(* Logix 5000 project; controller PLC_MCC1300_75F1 vendor 1 type 14 code 166 rev 32.11; software revision 32.04; part 29 of 83 *)
(* tags used below, declared in another part *)
   B3 : DINT[51];
   BENCH_BUZZER : ALIAS FOR O[74].12;
   C5 : COUNTER[51];
   CNV10_FLT : ALIAS FOR I[4].9;
   CNV11_FLT : ALIAS FOR I[4].10;
   CNV12_FLT : ALIAS FOR I[4].11;
   CNV1_FLT : ALIAS FOR I[4].0;
   CNV2_FLT : ALIAS FOR I[4].1;
   CNV3_FLT : ALIAS FOR I[4].2;
   CNV4_FLT : ALIAS FOR I[4].3;
   CNV5_FLT : ALIAS FOR I[4].4;
   CNV6_FLT : ALIAS FOR I[4].5;
   CNV7_FLT : ALIAS FOR I[4].6;
   CNV8_FLT : ALIAS FOR I[4].7;
   CNV9_FLT : ALIAS FOR I[4].8;
   CRUSH_ALL_ON : ALIAS FOR B3[0].0;
   DRV_STOP_DEB : ALIAS FOR T4[30].DN;
   FAST_BLINK : ALIAS FOR T4[2];
   Host_Read : INT[500];
   I : INT[128];   // Local Input Updates Input Slot 2
   M2_ALM_HORN_RLY : ALIAS FOR O[9].3;
   M2_BLUE_STKLTE : ALIAS FOR O[9].5;
   MMI_DATA : INT[64];   // MMI DATA For Fix 32
   MMI_FROM_MB : MESSAGE;
   MMI_TO_MB : MESSAGE;
   N130 : INT[8];
   N131 : INT[8];
   N14 : DINT[500];
   N72 : DINT[200];
   O : INT[128];
   REL_CRUSH_ALL_OFF : ALIAS FOR I[73].10;
   REL_CRUSH_ALL_ON : ALIAS FOR I[73].11;
   SLOW_BLINK : ALIAS FOR T4[0];
   T4 : TIMER[51];
   TD_ALM_HORN_RLY : ALIAS FOR O[21].3;
   TD_CS2S_Crush_All_Stacklight : ALIAS FOR O[70].15;   // Red Light mounted on the top of panel
   TD_DRV_FLT_LMP : ALIAS FOR O[21].0;
   TDN_CRUSH_ALL_OFF : ALIAS FOR I[44].12;
   TDN_CRUSH_ALL_ON : ALIAS FOR I[44].13;
   TDN_FLT : ALIAS FOR I[18].1;
   TDS_CRUSH_ALL_OFF : ALIAS FOR I[64].12;
   TDS_CRUSH_ALL_ON : ALIAS FOR I[64].13;
   TDS_FLT : ALIAS FOR I[18].2;
   TK_FLT : ALIAS FOR I[18].0;
   TMR_Power_Cycle : TIMER;
   xAlwaysOFF : BOOL;
(* MainProgram, continued *)

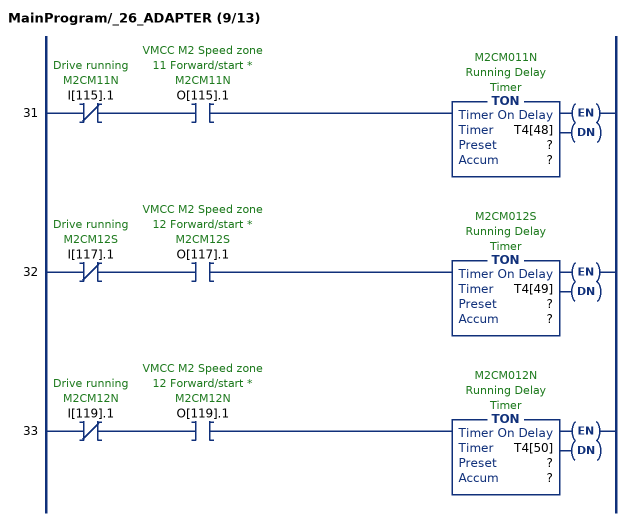
   31: XIO(I[115].1)XIC(O[115].1)TON(T4[48],?,?);
   32: XIO(I[117].1)XIC(O[117].1)TON(T4[49],?,?);
   33: XIO(I[119].1)XIC(O[119].1)TON(T4[50],?,?);
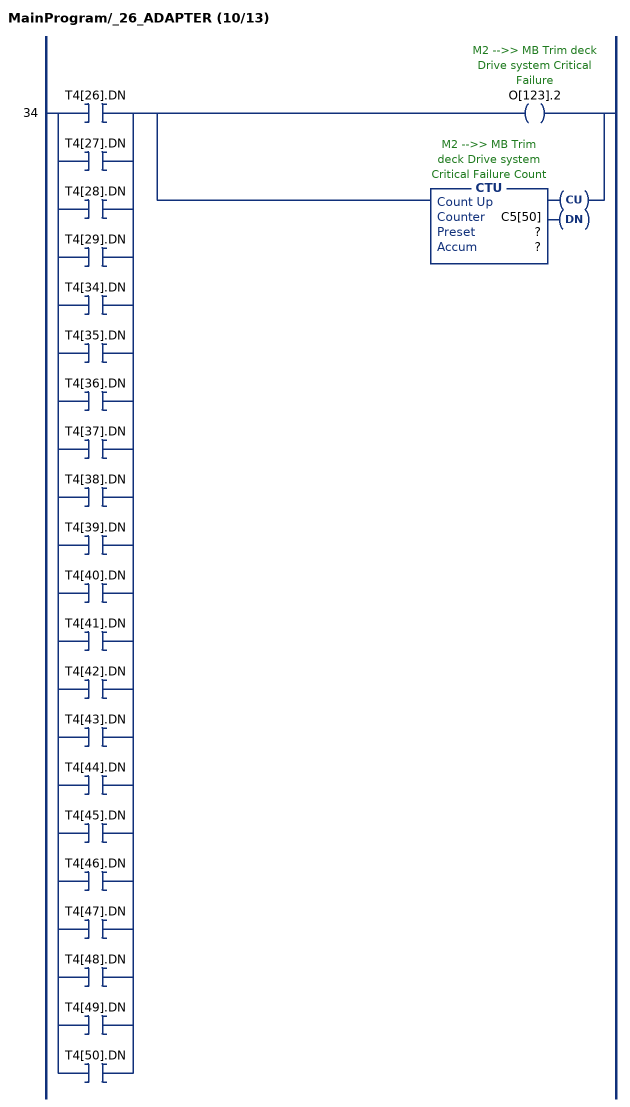
   34: [XIC(T4[26].DN) ,XIC(T4[27].DN) ,XIC(T4[28].DN) ,XIC(T4[29].DN) ,XIC(T4[34].DN) ,XIC(T4[35].DN) ,XIC(T4[36].DN) ,XIC(T4[37].DN) ,XIC(T4[38].DN) ,XIC(T4[39].DN) ,XIC(T4[40].DN) ,XIC(T4[41].DN) ,XIC(T4[42].DN) ,XIC(T4[43].DN) ,XIC(T4[44].DN) ,XIC(T4[45].DN) ,XIC(T4[46].DN) ,XIC(T4[47].DN) ,XIC(T4[48].DN) ,XIC(T4[49].DN) ,XIC(T4[50].DN) ][OTE(O[123].2) ,CTU(C5[50],?,?) ];
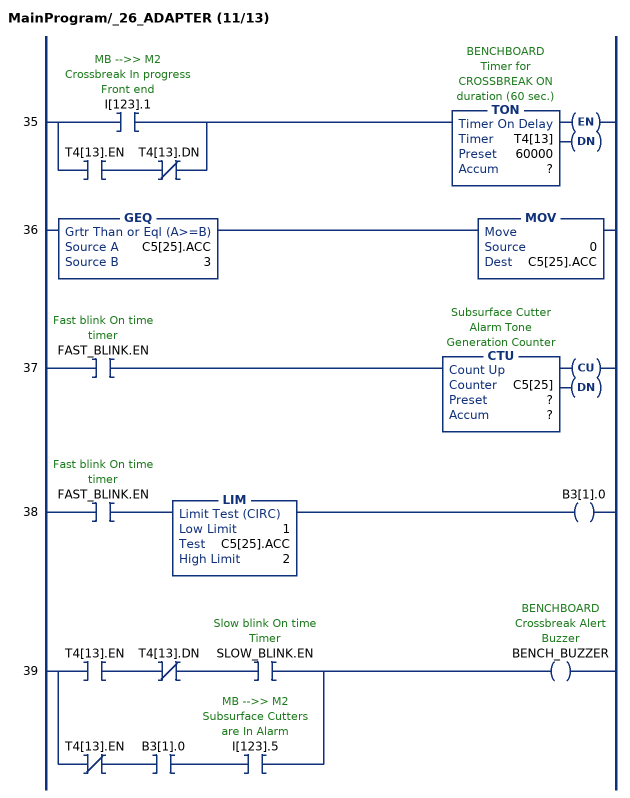
   35: [XIC(I[123].1) ,XIC(T4[13].EN) XIO(T4[13].DN) ]TON(T4[13],?,?);
   36: GEQ(C5[25].ACC,3)MOV(0,C5[25].ACC);
   37: XIC(FAST_BLINK.EN)CTU(C5[25],?,?);
   38: XIC(FAST_BLINK.EN)LIM(1,C5[25].ACC,2)OTE(B3[1].0);
   39: [XIC(T4[13].EN) XIO(T4[13].DN) XIC(SLOW_BLINK.EN) ,XIO(T4[13].EN) XIC(B3[1].0) XIC(I[123].5) ]OTE(BENCH_BUZZER);
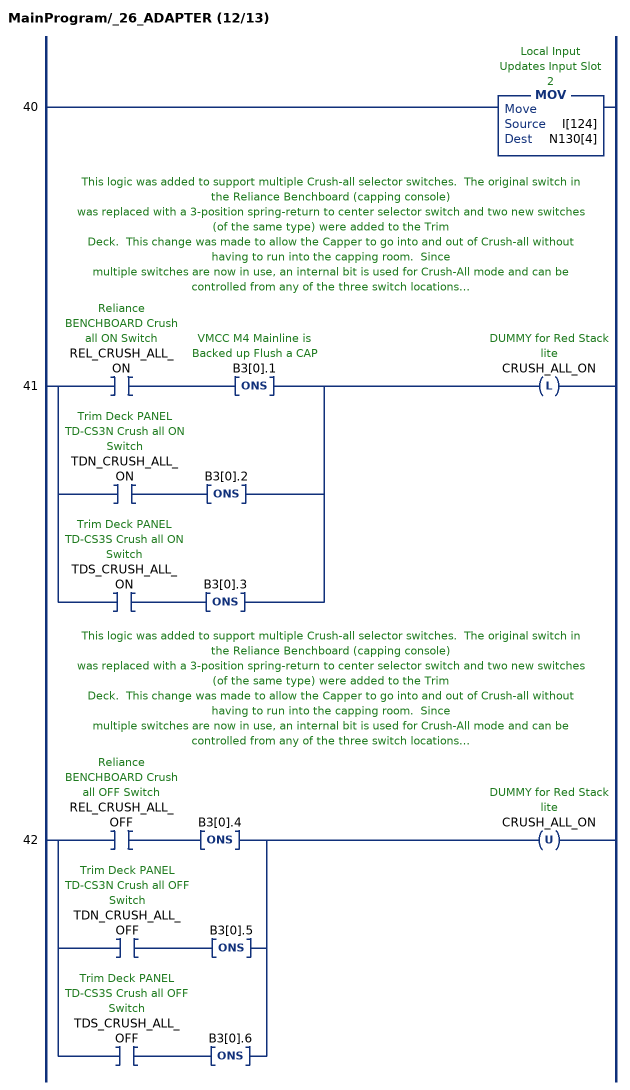
   40: MOV(I[124],N130[4]);
   // This logic was added to support multiple Crush-all selector switches.  The original switch in the Reliance Benchboard (capping console)
   // was replaced with a 3-position spring-return to center selector switch and two new switches (of the same type) were added to the Trim
   // Deck.  This change was made to allow the Capper to go into and out of Crush-all without having to run into the capping room.  Since
   // multiple switches are now in use, an internal bit is used for Crush-All mode and can be controlled from any of the three switch locations.
   // Note that one-shots [ONS] are used to keep a stuck-on selector switch contact from preventing the other two switches from operating
   // properly.  Also note that Latches and Unlatches are used (rather than a seal circuit) so that the system rides through power bumps properly
   // (i.e. Crush-all will stay in its current state, whether on or off, after a power bump).   DMK 10/21/02
   41: [XIC(REL_CRUSH_ALL_ON) ONS(B3[0].1) ,XIC(TDN_CRUSH_ALL_ON) ONS(B3[0].2) ,XIC(TDS_CRUSH_ALL_ON) ONS(B3[0].3) ]OTL(CRUSH_ALL_ON);
   // This logic was added to support multiple Crush-all selector switches.  The original switch in the Reliance Benchboard (capping console)
   // was replaced with a 3-position spring-return to center selector switch and two new switches (of the same type) were added to the Trim
   // Deck.  This change was made to allow the Capper to go into and out of Crush-all without having to run into the capping room.  Since
   // multiple switches are now in use, an internal bit is used for Crush-All mode and can be controlled from any of the three switch locations.
   // Note that one-shots [ONS] are used to keep a stuck-on selector switch contact from preventing the other two switches from operating
   // properly.  Also note that Latches and Unlatches are used (rather than a seal circuit) so that the system rides through power bumps properly
   // (i.e. Crush-all will stay in its current state, whether on or off, after a power bump).   DMK 10/21/02
   42: [XIC(REL_CRUSH_ALL_OFF) ONS(B3[0].4) ,XIC(TDN_CRUSH_ALL_OFF) ONS(B3[0].5) ,XIC(TDS_CRUSH_ALL_OFF) ONS(B3[0].6) ]OTU(CRUSH_ALL_ON);
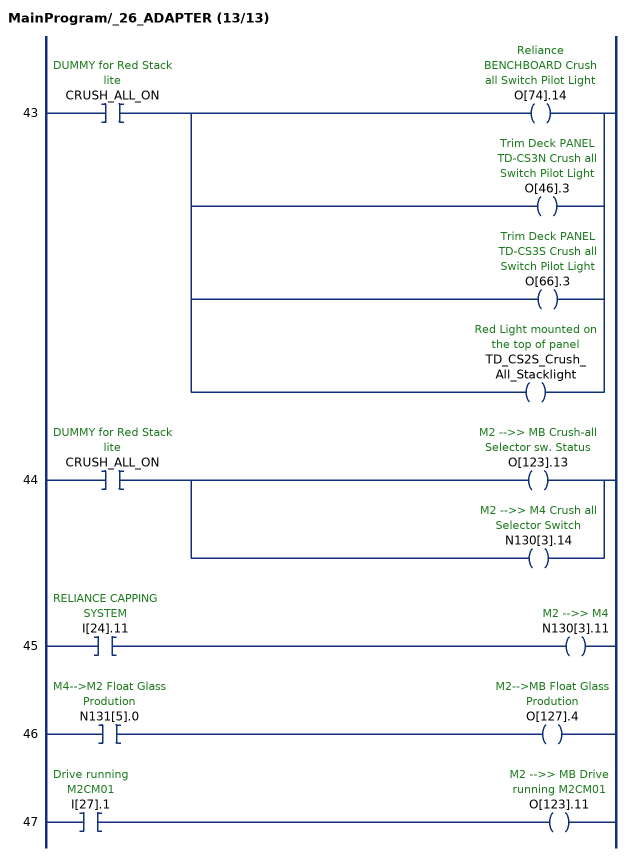
   43: XIC(CRUSH_ALL_ON)[OTE(O[74].14) ,OTE(O[46].3) ,OTE(O[66].3) ,OTE(TD_CS2S_Crush_All_Stacklight) ];
   44: XIC(CRUSH_ALL_ON)[OTE(O[123].13) ,OTE(N130[3].14) ];
   45: XIC(I[24].11)OTE(N130[3].11);
   46: XIC(N131[5].0)OTE(O[127].4);
   47: XIC(I[27].1)OTE(O[123].11);
END_ROUTINE

ROUTINE _2_MCP_A   (* ladder *)
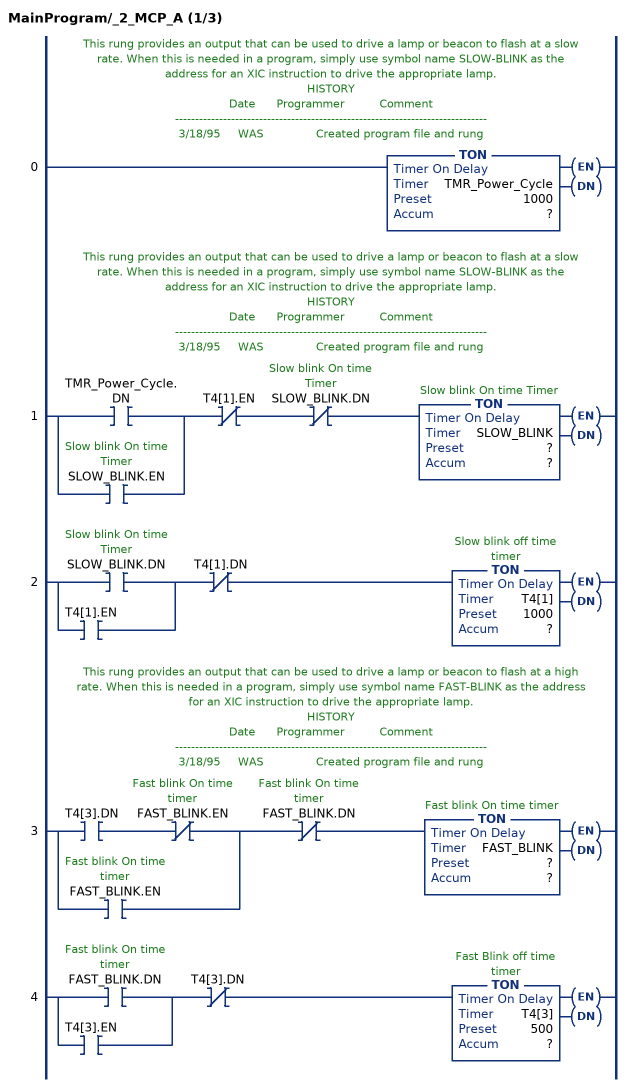
   // This rung provides an output that can be used to drive a lamp or beacon to flash at a slow rate. When this is needed in a program, simply use symbol name SLOW-BLINK as the address for an XIC instruction to drive the appropriate lamp.
   // HISTORY
   //             Date      Programmer          Comment
   // ------------------------------------------------------------------------------
   //             3/18/95     WAS               Created program file and rung
   0: TON(TMR_Power_Cycle,?,?);
   // This rung provides an output that can be used to drive a lamp or beacon to flash at a slow rate. When this is needed in a program, simply use symbol name SLOW-BLINK as the address for an XIC instruction to drive the appropriate lamp.
   // HISTORY
   //             Date      Programmer          Comment
   // ------------------------------------------------------------------------------
   //             3/18/95     WAS               Created program file and rung
   1: [XIC(TMR_Power_Cycle.DN) ,XIC(SLOW_BLINK.EN) ]XIO(T4[1].EN)XIO(SLOW_BLINK.DN)TON(SLOW_BLINK,?,?);
   2: [XIC(SLOW_BLINK.DN) ,XIC(T4[1].EN) ]XIO(T4[1].DN)TON(T4[1],?,?);
   // This rung provides an output that can be used to drive a lamp or beacon to flash at a high rate. When this is needed in a program, simply use symbol name FAST-BLINK as the address for an XIC instruction to drive the appropriate lamp.
   // HISTORY
   //             Date      Programmer          Comment
   // ------------------------------------------------------------------------------
   //             3/18/95     WAS               Created program file and rung
   3: [XIC(T4[3].DN) XIO(FAST_BLINK.EN) ,XIC(FAST_BLINK.EN) ]XIO(FAST_BLINK.DN)TON(FAST_BLINK,?,?);
   4: [XIC(FAST_BLINK.DN) ,XIC(T4[3].EN) ]XIO(T4[3].DN)TON(T4[3],?,?);
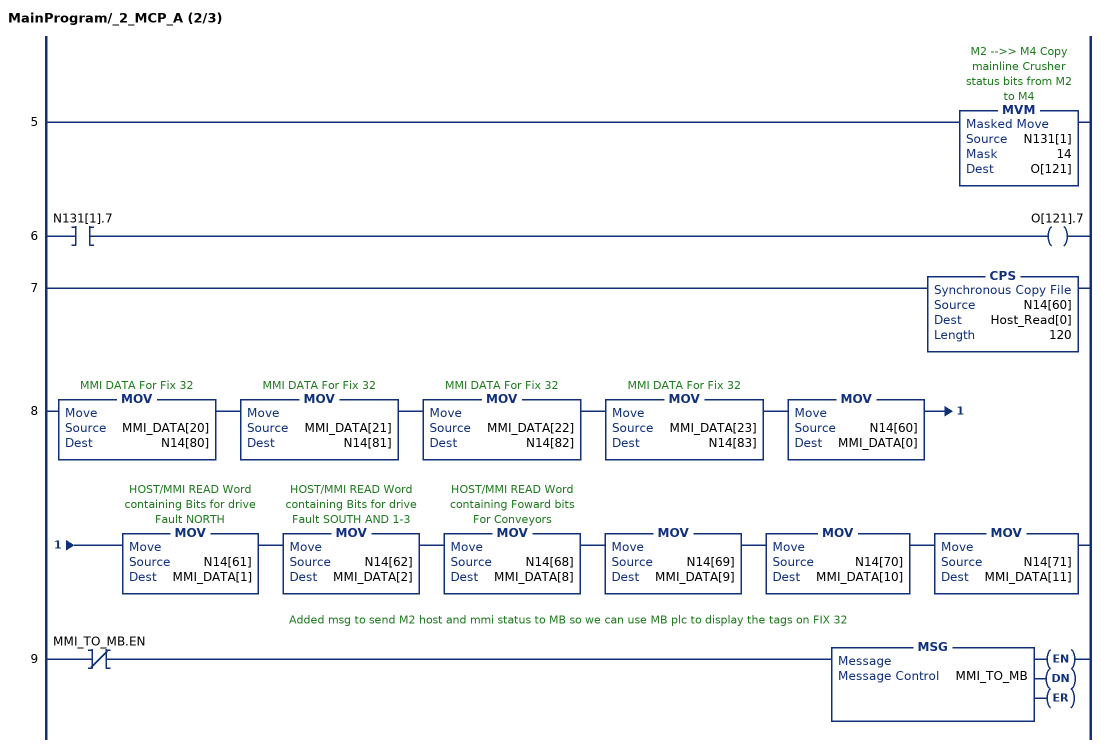
   5: MVM(N131[1],14,O[121]);
   6: XIC(N131[1].7)OTE(O[121].7);
   7: CPS(N14[60],Host_Read[0],120);
   8: MOV(MMI_DATA[20],N14[80])MOV(MMI_DATA[21],N14[81])MOV(MMI_DATA[22],N14[82])MOV(MMI_DATA[23],N14[83])MOV(N14[60],MMI_DATA[0])MOV(N14[61],MMI_DATA[1])MOV(N14[62],MMI_DATA[2])MOV(N14[68],MMI_DATA[8])MOV(N14[69],MMI_DATA[9])MOV(N14[70],MMI_DATA[10])MOV(N14[71],MMI_DATA[11]);
   // Added msg to send M2 host and mmi status to MB so we can use MB plc to display the tags on FIX 32
   9: XIO(MMI_TO_MB.EN)MSG(MMI_TO_MB);
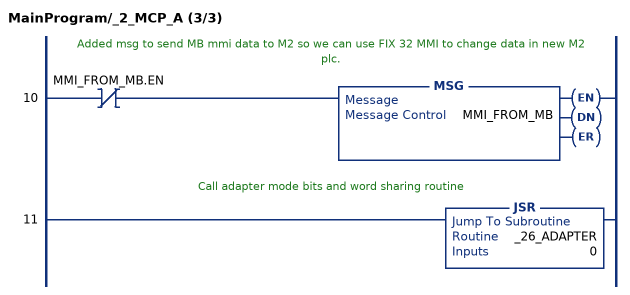
   // Added msg to send MB mmi data to M2 so we can use FIX 32 MMI to change data in new M2 plc.
   10: XIO(MMI_FROM_MB.EN)MSG(MMI_FROM_MB);
   // Call adapter mode bits and word sharing routine
   11: JSR(_26_ADAPTER,0);
END_ROUTINE

ROUTINE _3_MCP_B   (* ladder *)
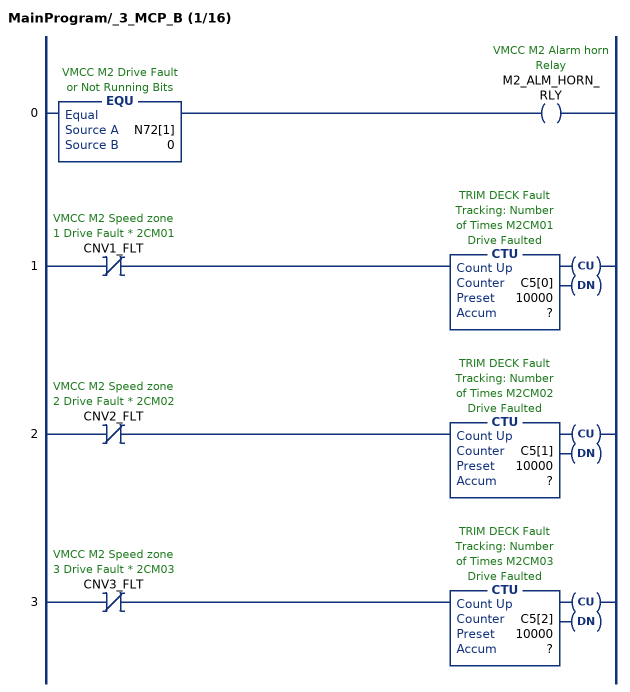
   0: EQU(N72[1],0)OTE(M2_ALM_HORN_RLY);
   1: XIO(CNV1_FLT)CTU(C5[0],?,?);
   2: XIO(CNV2_FLT)CTU(C5[1],?,?);
   3: XIO(CNV3_FLT)CTU(C5[2],?,?);
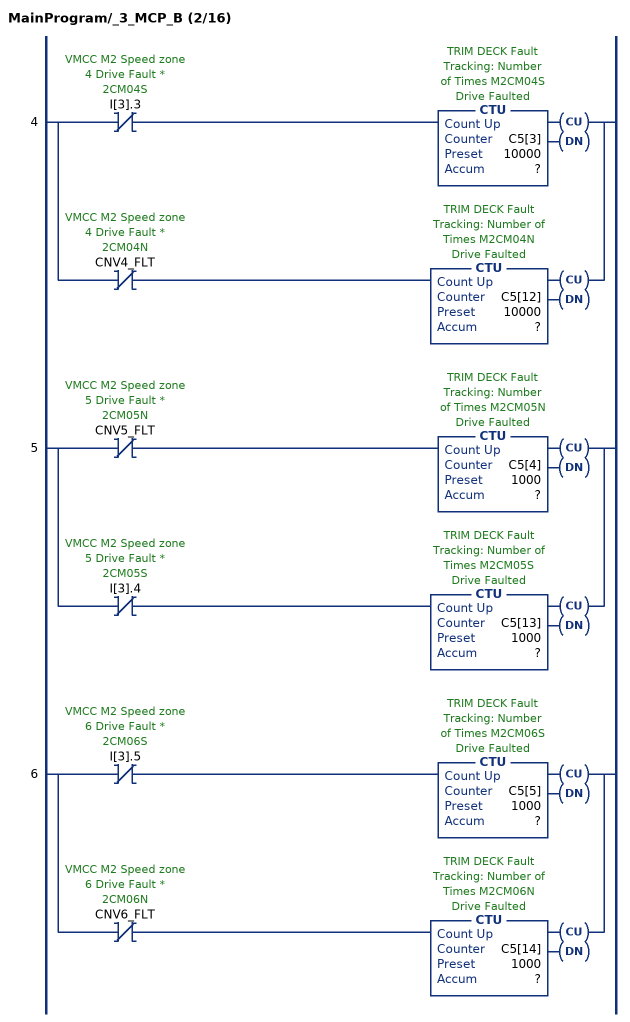
   4: [XIO(I[3].3) CTU(C5[3],?,?) ,XIO(CNV4_FLT) CTU(C5[12],?,?) ];
   5: [XIO(CNV5_FLT) CTU(C5[4],?,?) ,XIO(I[3].4) CTU(C5[13],?,?) ];
   6: [XIO(I[3].5) CTU(C5[5],?,?) ,XIO(CNV6_FLT) CTU(C5[14],?,?) ];
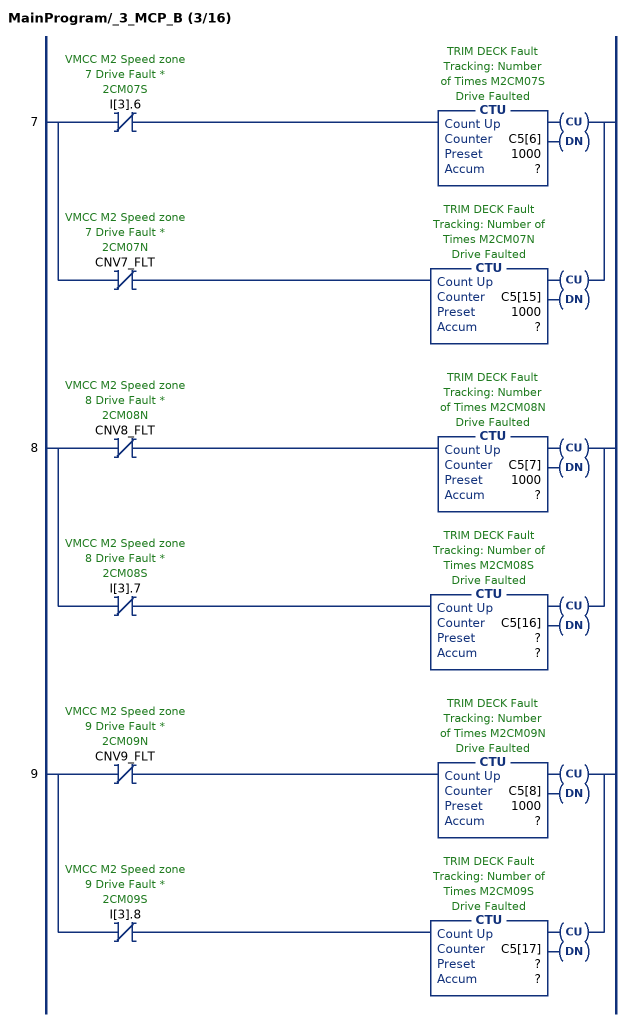
   7: [XIO(I[3].6) CTU(C5[6],?,?) ,XIO(CNV7_FLT) CTU(C5[15],?,?) ];
   8: [XIO(CNV8_FLT) CTU(C5[7],?,?) ,XIO(I[3].7) CTU(C5[16],?,?) ];
   9: [XIO(CNV9_FLT) CTU(C5[8],?,?) ,XIO(I[3].8) CTU(C5[17],?,?) ];
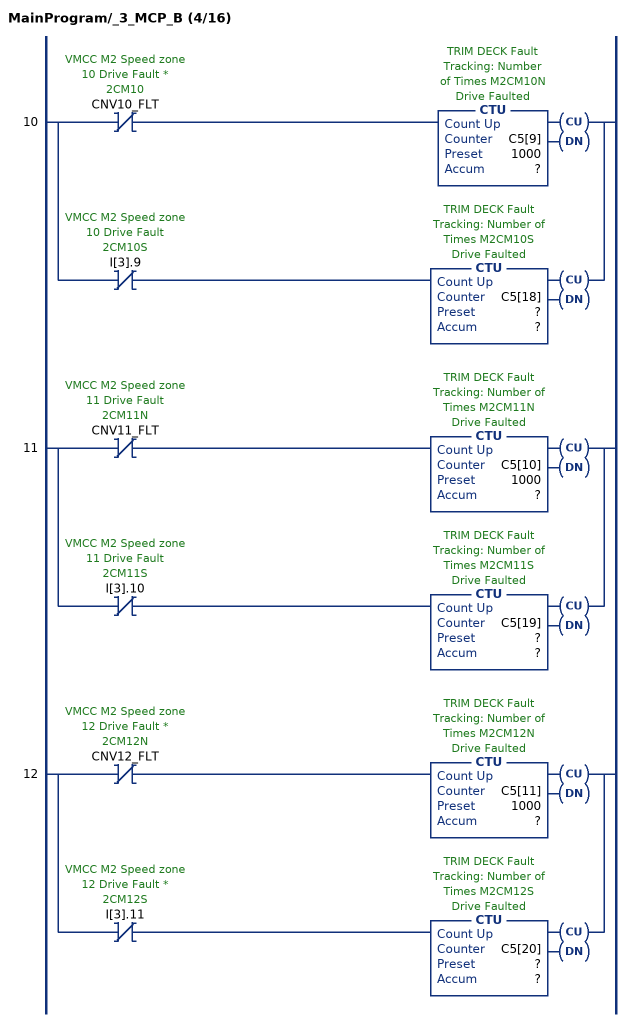
   10: [XIO(CNV10_FLT) CTU(C5[9],?,?) ,XIO(I[3].9) CTU(C5[18],?,?) ];
   11: [XIO(CNV11_FLT) CTU(C5[10],?,?) ,XIO(I[3].10) CTU(C5[19],?,?) ];
   12: [XIO(CNV12_FLT) CTU(C5[11],?,?) ,XIO(I[3].11) CTU(C5[20],?,?) ];
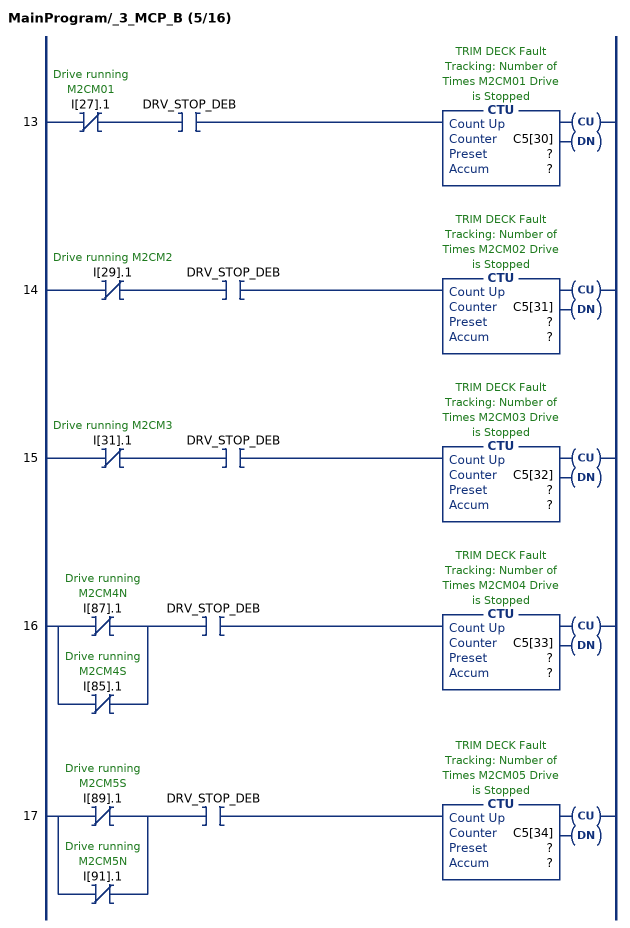
   13: XIO(I[27].1)XIC(DRV_STOP_DEB)CTU(C5[30],?,?);
   14: XIO(I[29].1)XIC(DRV_STOP_DEB)CTU(C5[31],?,?);
   15: XIO(I[31].1)XIC(DRV_STOP_DEB)CTU(C5[32],?,?);
   16: [XIO(I[87].1) ,XIO(I[85].1) ]XIC(DRV_STOP_DEB)CTU(C5[33],?,?);
   17: [XIO(I[89].1) ,XIO(I[91].1) ]XIC(DRV_STOP_DEB)CTU(C5[34],?,?);
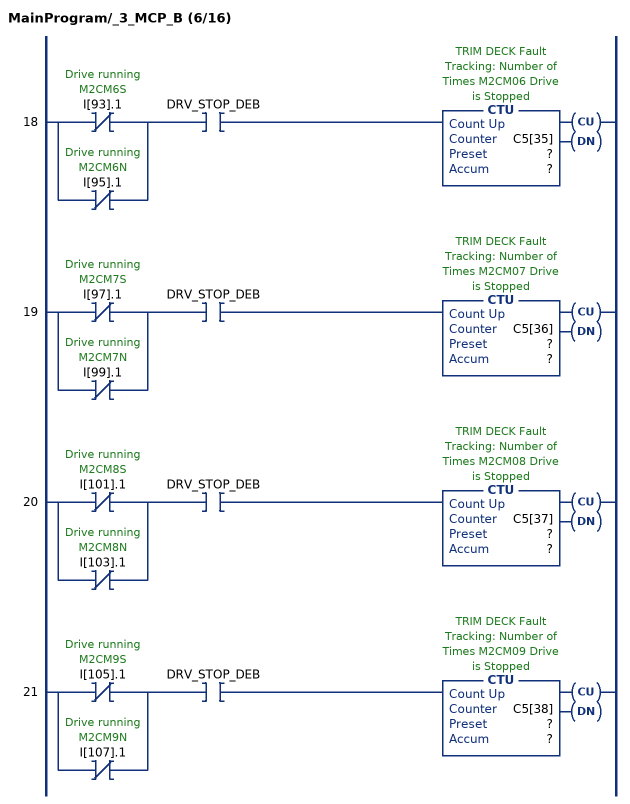
   18: [XIO(I[93].1) ,XIO(I[95].1) ]XIC(DRV_STOP_DEB)CTU(C5[35],?,?);
   19: [XIO(I[97].1) ,XIO(I[99].1) ]XIC(DRV_STOP_DEB)CTU(C5[36],?,?);
   20: [XIO(I[101].1) ,XIO(I[103].1) ]XIC(DRV_STOP_DEB)CTU(C5[37],?,?);
   21: [XIO(I[105].1) ,XIO(I[107].1) ]XIC(DRV_STOP_DEB)CTU(C5[38],?,?);
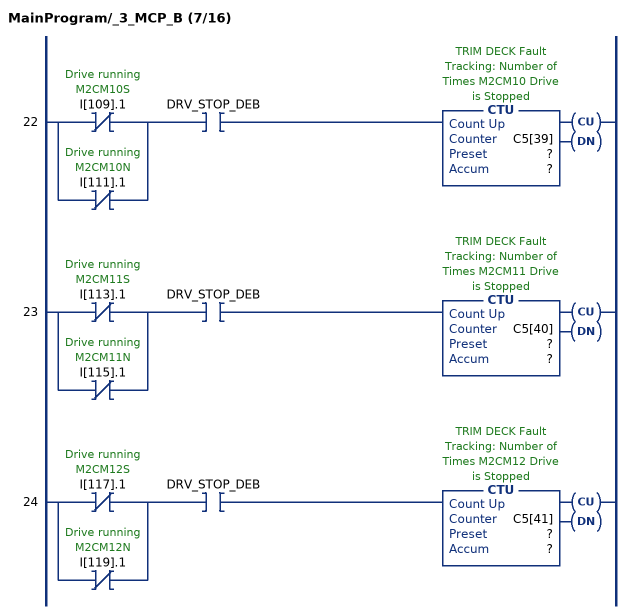
   22: [XIO(I[109].1) ,XIO(I[111].1) ]XIC(DRV_STOP_DEB)CTU(C5[39],?,?);
   23: [XIO(I[113].1) ,XIO(I[115].1) ]XIC(DRV_STOP_DEB)CTU(C5[40],?,?);
   24: [XIO(I[117].1) ,XIO(I[119].1) ]XIC(DRV_STOP_DEB)CTU(C5[41],?,?);
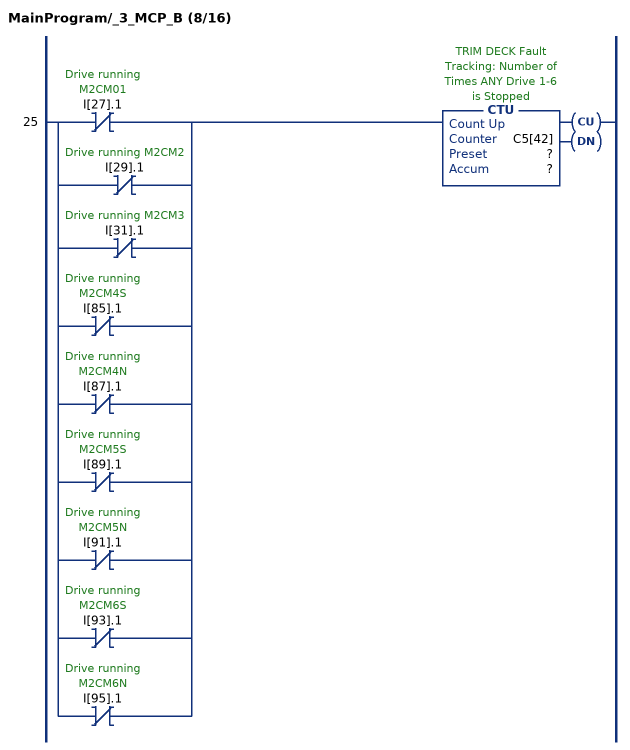
   25: [XIO(I[27].1) ,XIO(I[29].1) ,XIO(I[31].1) ,XIO(I[85].1) ,XIO(I[87].1) ,XIO(I[89].1) ,XIO(I[91].1) ,XIO(I[93].1) ,XIO(I[95].1) ]CTU(C5[42],?,?);
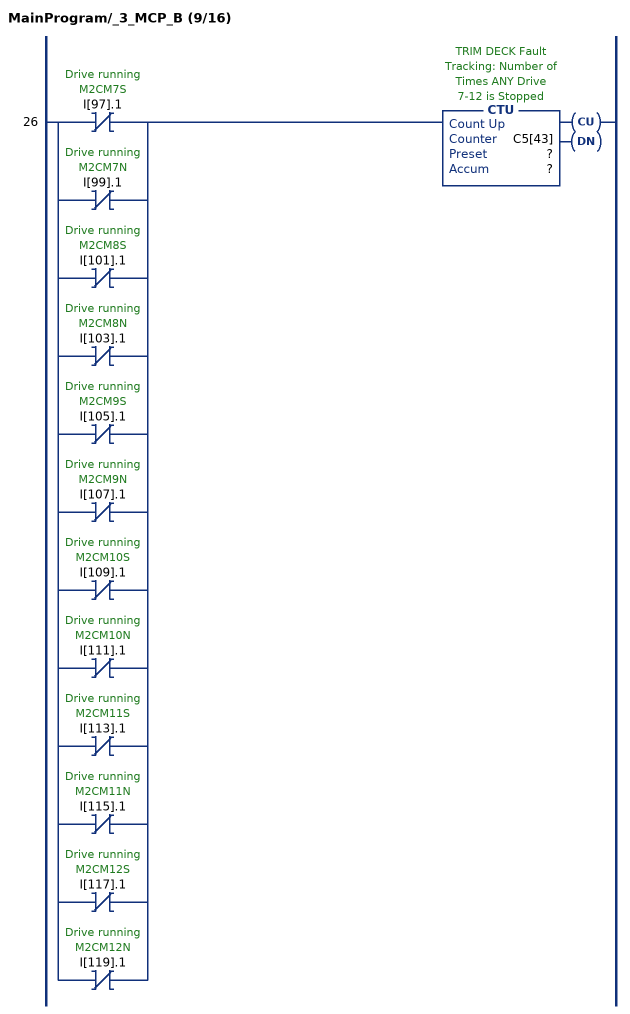
   26: [XIO(I[97].1) ,XIO(I[99].1) ,XIO(I[101].1) ,XIO(I[103].1) ,XIO(I[105].1) ,XIO(I[107].1) ,XIO(I[109].1) ,XIO(I[111].1) ,XIO(I[113].1) ,XIO(I[115].1) ,XIO(I[117].1) ,XIO(I[119].1) ]CTU(C5[43],?,?);
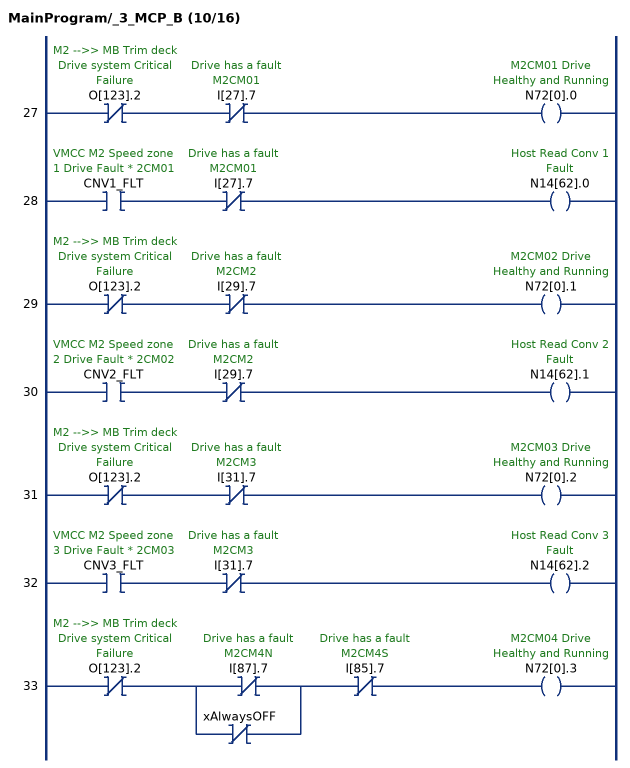
   27: XIO(O[123].2)XIO(I[27].7)OTE(N72[0].0);
   28: XIC(CNV1_FLT)XIO(I[27].7)OTE(N14[62].0);
   29: XIO(O[123].2)XIO(I[29].7)OTE(N72[0].1);
   30: XIC(CNV2_FLT)XIO(I[29].7)OTE(N14[62].1);
   31: XIO(O[123].2)XIO(I[31].7)OTE(N72[0].2);
   32: XIC(CNV3_FLT)XIO(I[31].7)OTE(N14[62].2);
   33: XIO(O[123].2)[XIO(I[87].7) ,XIO(xAlwaysOFF) ]XIO(I[85].7)OTE(N72[0].3);
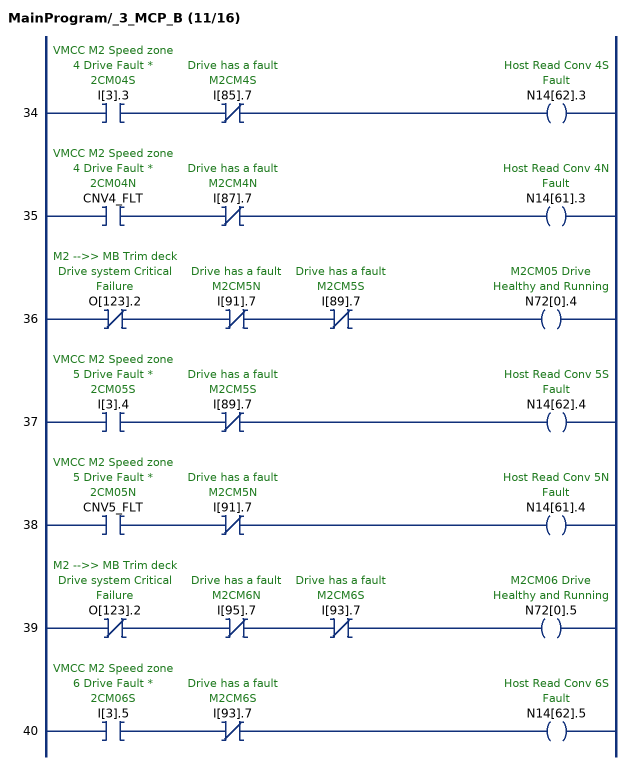
   34: XIC(I[3].3)XIO(I[85].7)OTE(N14[62].3);
   35: XIC(CNV4_FLT)XIO(I[87].7)OTE(N14[61].3);
   36: XIO(O[123].2)XIO(I[91].7)XIO(I[89].7)OTE(N72[0].4);
   37: XIC(I[3].4)XIO(I[89].7)OTE(N14[62].4);
   38: XIC(CNV5_FLT)XIO(I[91].7)OTE(N14[61].4);
   39: XIO(O[123].2)XIO(I[95].7)XIO(I[93].7)OTE(N72[0].5);
   40: XIC(I[3].5)XIO(I[93].7)OTE(N14[62].5);
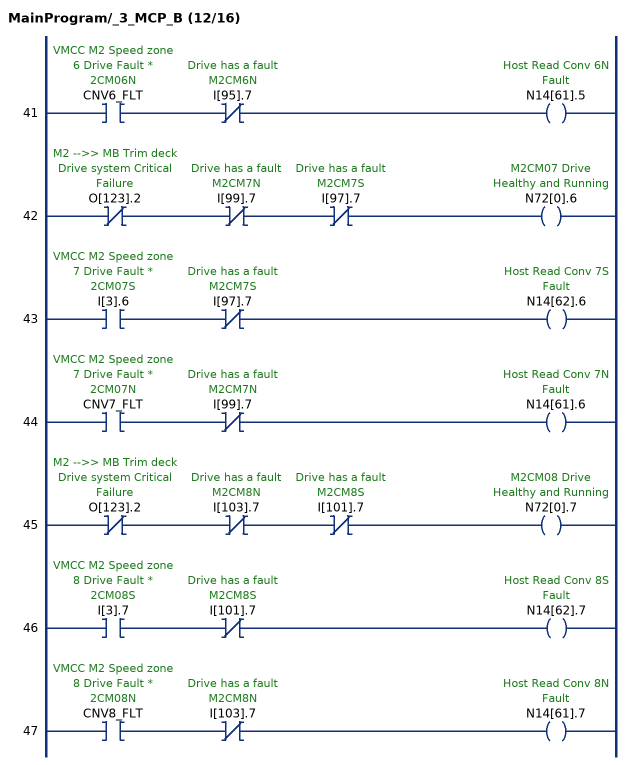
   41: XIC(CNV6_FLT)XIO(I[95].7)OTE(N14[61].5);
   42: XIO(O[123].2)XIO(I[99].7)XIO(I[97].7)OTE(N72[0].6);
   43: XIC(I[3].6)XIO(I[97].7)OTE(N14[62].6);
   44: XIC(CNV7_FLT)XIO(I[99].7)OTE(N14[61].6);
   45: XIO(O[123].2)XIO(I[103].7)XIO(I[101].7)OTE(N72[0].7);
   46: XIC(I[3].7)XIO(I[101].7)OTE(N14[62].7);
   47: XIC(CNV8_FLT)XIO(I[103].7)OTE(N14[61].7);
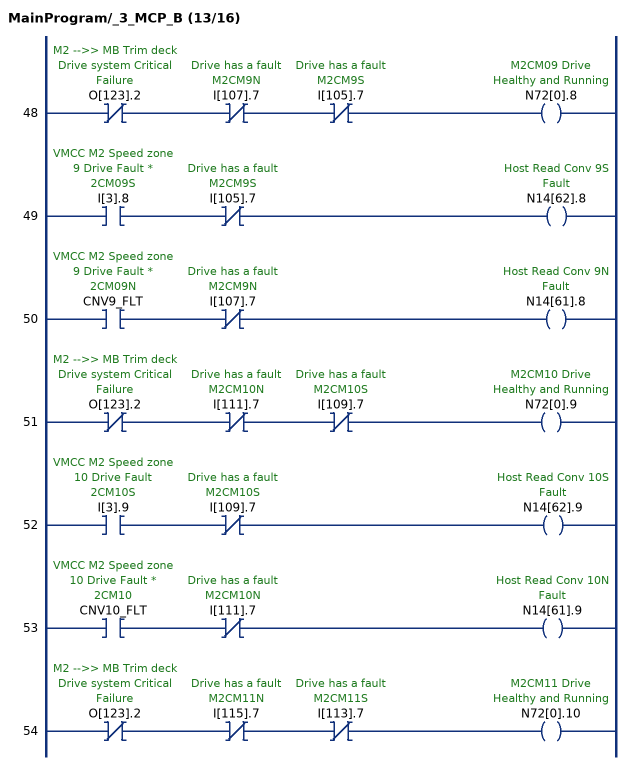
   48: XIO(O[123].2)XIO(I[107].7)XIO(I[105].7)OTE(N72[0].8);
   49: XIC(I[3].8)XIO(I[105].7)OTE(N14[62].8);
   50: XIC(CNV9_FLT)XIO(I[107].7)OTE(N14[61].8);
   51: XIO(O[123].2)XIO(I[111].7)XIO(I[109].7)OTE(N72[0].9);
   52: XIC(I[3].9)XIO(I[109].7)OTE(N14[62].9);
   53: XIC(CNV10_FLT)XIO(I[111].7)OTE(N14[61].9);
   54: XIO(O[123].2)XIO(I[115].7)XIO(I[113].7)OTE(N72[0].10);
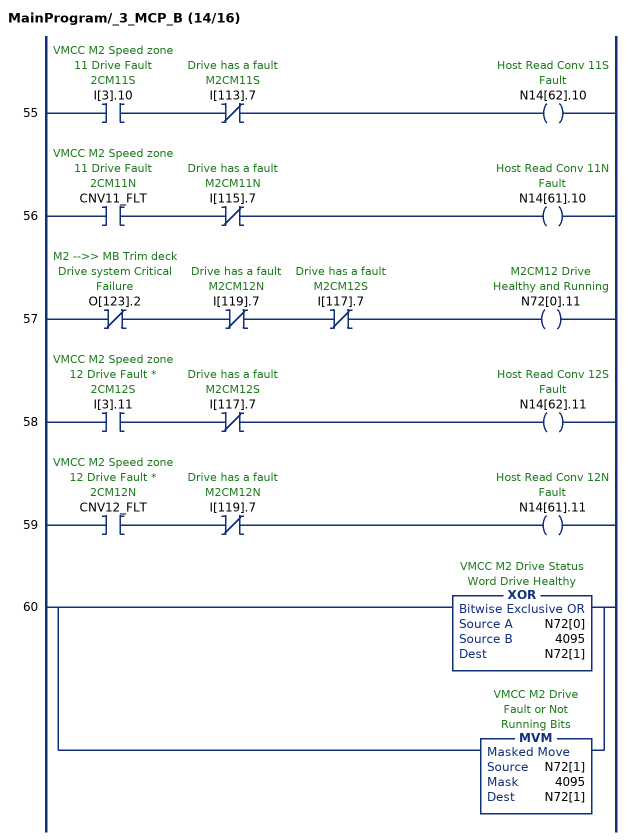
   55: XIC(I[3].10)XIO(I[113].7)OTE(N14[62].10);
   56: XIC(CNV11_FLT)XIO(I[115].7)OTE(N14[61].10);
   57: XIO(O[123].2)XIO(I[119].7)XIO(I[117].7)OTE(N72[0].11);
   58: XIC(I[3].11)XIO(I[117].7)OTE(N14[62].11);
   59: XIC(CNV12_FLT)XIO(I[119].7)OTE(N14[61].11);
   60: [XOR(N72[0],4095,N72[1]) ,MVM(N72[1],4095,N72[1]) ];
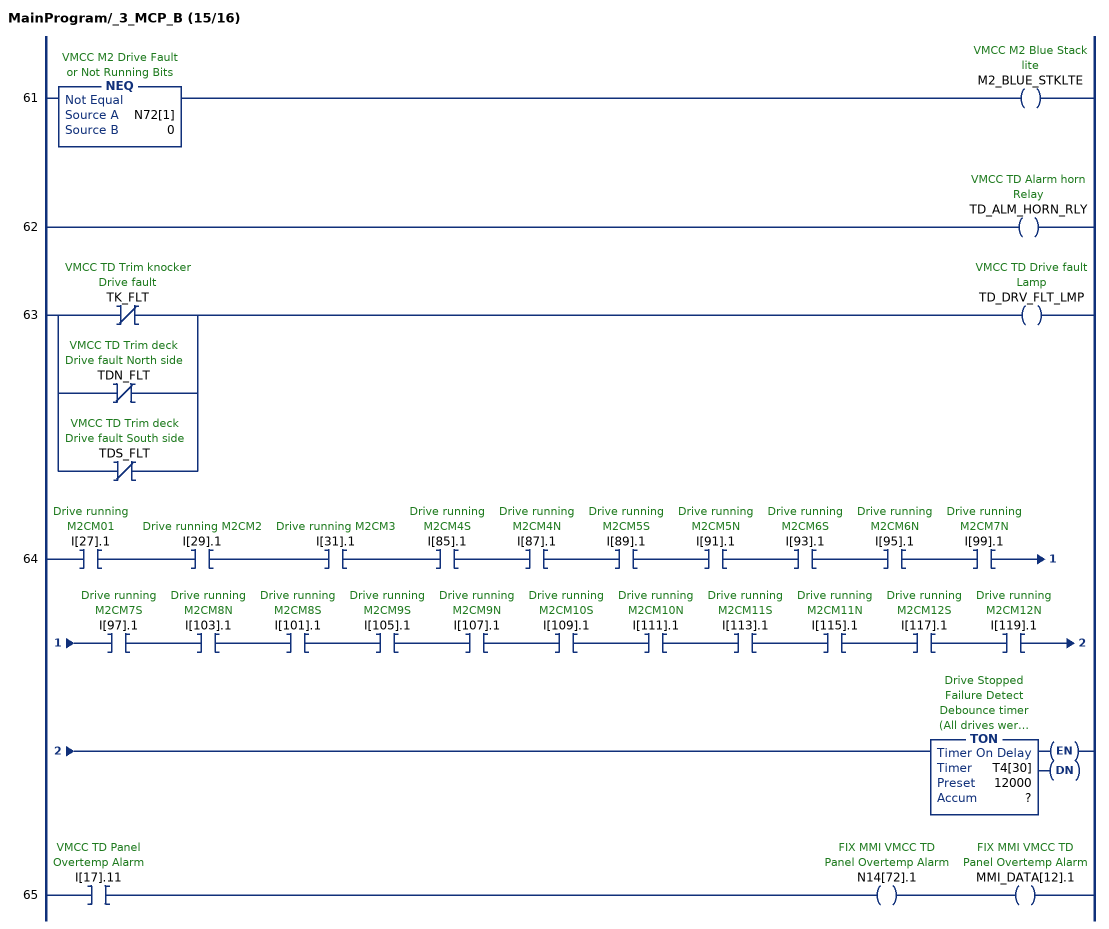
   61: NEQ(N72[1],0)OTE(M2_BLUE_STKLTE);
   62: OTE(TD_ALM_HORN_RLY);
   63: [XIO(TK_FLT) ,XIO(TDN_FLT) ,XIO(TDS_FLT) ]OTE(TD_DRV_FLT_LMP);
   64: XIC(I[27].1)XIC(I[29].1)XIC(I[31].1)XIC(I[85].1)XIC(I[87].1)XIC(I[89].1)XIC(I[91].1)XIC(I[93].1)XIC(I[95].1)XIC(I[99].1)XIC(I[97].1)XIC(I[103].1)XIC(I[101].1)XIC(I[105].1)XIC(I[107].1)XIC(I[109].1)XIC(I[111].1)XIC(I[113].1)XIC(I[115].1)XIC(I[117].1)XIC(I[119].1)TON(T4[30],?,?);
   65: XIC(I[17].11)OTE(N14[72].1)OTE(MMI_DATA[12].1);
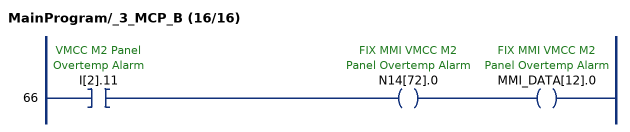
   66: XIC(I[2].11)OTE(N14[72].0)OTE(MMI_DATA[12].0);
END_ROUTINE
